(* Logix 5000 project; controller FV vendor 1 type 14 code 217 rev 31.11; software revision 31.00; part 2 of 63 *)

        [144]   // 0 0 0 min input
        [145]   // 0 0 0 max input
        [146]   // 0 0 0 min scaled
        [147]   // 0 0 0 max scale
        [148]   // 0 0 0 High Limit
        [149]   // 0 0 0 Low Limit
        [14]   // FV26/LTX01 FV26 level transmitter min input
        [151]   // 0 0 0 Flags
        [151].0   // 0 0 0 High
        [151].1   // 0 0 0 Low
        [151].15   // 0 0 0 Fault
        [152]   // 0 0 0 mA
        [153]   // 0 0 0 spare
        [154]   // 0 0 0 min input
        [155]   // 0 0 0 max input
        [156]   // 0 0 0 min scaled
        [157]   // 0 0 0 max scale
        [158]   // 0 0 0 High Limit
        [159]   // 0 0 0 Low Limit
        [15]   // FV26/LTX01 FV26 level transmitter max input
        [16]   // FV26/LTX01 FV26 level transmitter min scaled
        [17]   // FV26/LTX01 FV26 level transmitter max scale
        [18]   // FV26/LTX01 FV26 level transmitter High Limit
        [19]   // FV26/LTX01 FV26 level transmitter Low Limit
        [1]   // FV26/PTX01 FV26 top pressure Flags
        [1].0   // FV26/PTX01 FV26 top pressure High
        [1].1   // FV26/PTX01 FV26 top pressure Low
        [1].15   // FV26/PTX01 FV26 top pressure Fault
        [20]   // FV27/PTX01 FV27 top pressure transmitter
        [21]   // FV27/PTX01 FV27 top pressure Flags
        [21].0   // FV27/PTX01 FV27 top pressure High
        [21].1   // FV27/PTX01 FV27 top pressure Low
        [21].15   // FV27/PTX01 FV27 top pressure Fault
        [22]   // FV27/PTX01 FV27 top pressure mA
        [23]   // FV27/PTX01 FV27 top pressure spare
        [24]   // FV27/PTX01 FV27 top pressure min input
        [25]   // FV27/PTX01 FV27 top pressure max input
        [26]   // FV27/PTX01 FV27 top pressure min scaled
        [27]   // FV27/PTX01 FV27 top pressure max scale
        [28]   // FV27/PTX01 FV27 top pressure High Limit
        [29]   // FV27/PTX01 FV27 top pressure Low Limit
        [2]   // FV26/PTX01 FV26 top pressure mA
        [30]   // FV27/LTX01 FV27 level transmitter
        [31]   // FV27/LTX01 FV27 level transmitter Flags
        [31].0   // FV27/LTX01 FV27 level transmitter High
        [31].1   // FV27/LTX01 FV27 level transmitter Low
        [31].15   // FV27/LTX01 FV27 level transmitter Fault
        [32]   // FV27/LTX01 FV27 level transmitter mA
        [33]   // FV27/LTX01 FV27 level transmitter spare
        [34]   // FV27/LTX01 FV27 level transmitter min input
        [35]   // FV27/LTX01 FV27 level transmitter max input
        [36]   // FV27/LTX01 FV27 level transmitter min scaled
        [37]   // FV27/LTX01 FV27 level transmitter max scale
        [38]   // FV27/LTX01 FV27 level transmitter High Limit
        [39]   // FV27/LTX01 FV27 level transmitter Low Limit
        [3]   // FV26/PTX01 FV26 top pressure spare
        [40]   // FV28/PTX01 FV28 top pressure transmitter
        [41]   // FV28/PTX01 FV28 top pressure Flags
        [41].0   // FV28/PTX01 FV28 top pressure High
        [41].1   // FV28/PTX01 FV28 top pressure Low
        [41].15   // FV28/PTX01 FV28 top pressure Fault
        [42]   // FV28/PTX01 FV28 top pressure mA
        [43]   // FV28/PTX01 FV28 top pressure spare
        [44]   // FV28/PTX01 FV28 top pressure min input
        [45]   // FV28/PTX01 FV28 top pressure max input
        [46]   // FV28/PTX01 FV28 top pressure min scaled
        [47]   // FV28/PTX01 FV28 top pressure max scale
        [48]   // FV28/PTX01 FV28 top pressure High Limit
        [49]   // FV28/PTX01 FV28 top pressure Low Limit
        [4]   // FV26/PTX01 FV26 top pressure min input
        [50]   // FV28/LTX01 FV28 level transmitter
        [51]   // FV28/LTX01 FV28 level transmitter Flags
        [51].0   // FV28/LTX01 FV28 level transmitter High
        [51].1   // FV28/LTX01 FV28 level transmitter Low
        [51].15   // FV28/LTX01 FV28 level transmitter Fault
        [52]   // FV28/LTX01 FV28 level transmitter mA
        [53]   // FV28/LTX01 FV28 level transmitter spare
        [54]   // FV28/LTX01 FV28 level transmitter min input
        [55]   // FV28/LTX01 FV28 level transmitter max input
        [56]   // FV28/LTX01 FV28 level transmitter min scaled
        [57]   // FV28/LTX01 FV28 level transmitter max scale
        [58]   // FV28/LTX01 FV28 level transmitter High Limit
        [59]   // FV28/LTX01 FV28 level transmitter Low Limit
        [5]   // FV26/PTX01 FV26 top pressure max input
        [60]   // FV29/PTX01 FV29 top pressure transmitter
        [61]   // FV29/PTX01 FV29 top pressure Flags
        [61].0   // FV29/PTX01 FV29 top pressure High
        [61].1   // FV29/PTX01 FV29 top pressure Low
        [61].15   // FV29/PTX01 FV29 top pressure Fault
        [62]   // FV29/PTX01 FV29 top pressure mA
        [63]   // FV29/PTX01 FV29 top pressure spare
        [64]   // FV29/PTX01 FV29 top pressure min input
        [65]   // FV29/PTX01 FV29 top pressure max input
        [66]   // FV29/PTX01 FV29 top pressure min scaled
        [67]   // FV29/PTX01 FV29 top pressure max scale
        [68]   // FV29/PTX01 FV29 top pressure High Limit
        [69]   // FV29/PTX01 FV29 top pressure Low Limit
        [6]   // FV26/PTX01 FV26 top pressure min scaled
        [70]   // FV29/LTX01 FV29 level transmitter
        [71]   // FV29/LTX01 FV29 level transmitter Flags
        [71].0   // FV29/LTX01 FV29 level transmitter High
        [71].1   // FV29/LTX01 FV29 level transmitter Low
        [71].15   // FV29/LTX01 FV29 level transmitter Fault
        [72]   // FV29/LTX01 FV29 level transmitter mA
        [73]   // FV29/LTX01 FV29 level transmitter spare
        [74]   // FV29/LTX01 FV29 level transmitter min input
        [75]   // FV29/LTX01 FV29 level transmitter max input
        [76]   // FV29/LTX01 FV29 level transmitter min scaled
        [77]   // FV29/LTX01 FV29 level transmitter max scale
        [78]   // FV29/LTX01 FV29 level transmitter High Limit
        [79]   // FV29/LTX01 FV29 level transmitter Low Limit
        [7]   // FV26/PTX01 FV26 top pressure max scale
        [80]   // FV30/PTX01 FV30 top pressure transmitter
        [81]   // FV30/PTX01 FV30 top pressure Flags
        [81].0   // FV30/PTX01 FV30 top pressure High
        [81].1   // FV30/PTX01 FV30 top pressure Low
        [81].15   // FV30/PTX01 FV30 top pressure Fault
        [82]   // FV30/PTX01 FV30 top pressure mA
        [83]   // FV30/PTX01 FV30 top pressure spare
        [84]   // FV30/PTX01 FV30 top pressure min input
        [85]   // FV30/PTX01 FV30 top pressure max input
        [86]   // FV30/PTX01 FV30 top pressure min scaled
        [87]   // FV30/PTX01 FV30 top pressure max scale
        [88]   // FV30/PTX01 FV30 top pressure High Limit
        [89]   // FV30/PTX01 FV30 top pressure Low Limit
        [8]   // FV26/PTX01 FV26 top pressure High Limit
        [90]   // FV30/LTX01 FV30 level transmitter
        [91]   // FV30/LTX01 FV30 level transmitter Flags
        [91].0   // FV30/LTX01 FV30 level transmitter High
        [91].1   // FV30/LTX01 FV30 level transmitter Low
        [91].15   // FV30/LTX01 FV30 level transmitter Fault
        [92]   // FV30/LTX01 FV30 level transmitter mA
        [93]   // FV30/LTX01 FV30 level transmitter spare
        [94]   // FV30/LTX01 FV30 level transmitter min input
        [95]   // FV30/LTX01 FV30 level transmitter max input
        [96]   // FV30/LTX01 FV30 level transmitter min scaled
        [97]   // FV30/LTX01 FV30 level transmitter max scale
        [98]   // FV30/LTX01 FV30 level transmitter High Limit
        [99]   // FV30/LTX01 FV30 level transmitter Low Limit
        [9]   // FV26/PTX01 FV26 top pressure Low Limit
   FR_N201 : INT[265];   // Original N File From SLC, No Description Available
   FR_N207 : INT[265] := ([0] := 256, [1] := 1, [2] := 2, [3] := 3, [4] := 4, [5] := 5, [6] := 6, [7] := 7, [8] := 8, [9] := 9, [10] := 10, [11] := 11, [12] := 12, [13] := 13, [14] := 14, [15] := 15, [16] := 16, [17] := 17, [18] := 18, [19] := 19, [20] := 20, [21] := 21, [22] := 22, [23] := 23, [24] := 24, [25] := 25, [26] := 26, [27] := 27, [28] := 28, [29] := 29, [30] := 30, [31] := 31, [32] := 32, [33] := 33, [34] := 34, [35] := 35, [36] := 36, [37] := 37, [38] := 38, [39] := 39, [40] := 40, [41] := 41, [42] := 42, [43] := 43, [44] := 44, [45] := 45, [46] := 46, [47] := 47, [48] := 48, [49] := 49, [50] := 50, [51] := 51, [52] := 52, [53] := 53, [54] := 54, [55] := 55, [56] := 56, [57] := 57, [58] := 58, [59] := 59,
        [60] := 60, [61] := 61, [62] := 62, [63] := 63, [64] := 64, [65] := 65, [66] := 66, [67] := 67, [68] := 68, [69] := 69, [70] := 70, [71] := 71, [72] := 72, [73] := 73, [74] := 74, [75] := 75, [76] := 76, [77] := 77, [78] := 78, [79] := 79, [80] := 80, [81] := 81, [82] := 82, [83] := 83, [84] := 84, [85] := 85, [86] := 86, [87] := 87, [88] := 88, [89] := 89, [90] := 90, [91] := 91, [92] := 92, [93] := 93, [94] := 94, [95] := 95, [96] := 96, [97] := 97, [98] := 98, [99] := 99, [100] := 100, [101] := 101, [102] := 102, [103] := 103, [104] := 104, [105] := 105, [106] := 106, [107] := 107, [108] := 108, [109] := 109, [110] := 110, [111] := 111, [112] := 112, [113] := 113, [114] := 114, [115] := 115, [116] := 116, [117] := 117, [118] := 118, [119] := 119,
        [120] := 120, [121] := 121, [122] := 122, [123] := 123, [124] := 124, [125] := 125, [126] := 126, [127] := 127, [128] := 128, [129] := 129, [130] := 130, [131] := 131, [132] := 132, [133] := 133, [134] := 134, [135] := 135, [136] := 136, [137] := 137, [138] := 138, [139] := 139, [140] := 140, [141] := 141, [142] := 142, [143] := 143, [144] := 144, [145] := 145, [146] := 146, [147] := 147, [148] := 148, [149] := 149, [150] := 150, [151] := 151, [152] := 152, [153] := 153, [154] := 154, [155] := 155, [156] := 156, [157] := 157, [158] := 158, [159] := 159, [160] := 160, [161] := 161, [162] := 162, [163] := 163, [164] := 164, [165] := 165, [166] := 166, [167] := 167, [168] := 168, [169] := 169, [170] := 170, [171] := 171, [172] := 172, [173] := 173, [174] := 174, [175] := 175, [176] := 176, [177] := 177, [178] := 178, [179] := 179,
        [180] := 180, [181] := 181, [182] := 182, [183] := 183, [184] := 184, [185] := 185, [186] := 186, [187] := 187, [188] := 188, [189] := 189, [190] := 190, [191] := 191, [192] := 192, [193] := 193, [194] := 194, [195] := 195, [196] := 196, [197] := 197, [198] := 198, [199] := 199, [200] := 200, [201] := 201, [202] := 202, [203] := 203, [204] := 204, [205] := 205, [206] := 206, [207] := 207, [208] := 208, [209] := 209, [210] := 210, [211] := 211, [212] := 212, [213] := 213, [214] := 214, [215] := 215, [216] := 216, [217] := 217, [218] := 218, [219] := 219, [220] := 220, [221] := 221, [222] := 222, [223] := 223, [224] := 224, [225] := 225, [226] := 226, [227] := 227, [228] := 228, [229] := 229, [230] := 230, [231] := 231, [232] := 232, [233] := 233, [234] := 234, [235] := 235, [236] := 236, [237] := 237, [238] := 238, [239] := 239,
        [240] := 240, [241] := 241, [242] := 242, [243] := 243, [244] := 244, [245] := 245, [246] := 246, [247] := 247, [248] := 248, [249] := 249, [250] := 250, [251] := 251, [252] := 252, [253] := 253, [254] := 254, [255] := 255);   // Original N File From SLC, No Description Available
   FR_N21 : INT[265] := ([26] := 700, [27] := 700, [28] := 700, [29] := 700, [30] := 700, [31] := 700);   // CHASE_V FV Filling Beer Chas e Volumes
   FR_N210 : INT[265] := ([0] := 500, [1] := 12000, [2] := 18725, [5] := 1000, [6] := 4000, [7] := 20000, [8] := 6242, [9] := 31208, [11] := 12000, [12] := 18725, [15] := 1000, [16] := 4000, [17] := 20000, [18] := 6242, [19] := 31208, [20] := 500, [21] := 8800, [22] := 13732, [25] := 1000, [26] := 4000, [27] := 20000, [28] := 6242, [29] := 31208);   // ANALOG_OUT Analog Outputs
        [0]   // YM/P01 Yeast Main Pump 1 FV26-31 0.0-100.0%
        [10]   // YM/P02 Yeast Main Pump 2 FV1-17 0.0-100.0%
        [11]   // YM/P02 Yeast Main Pump 2 FV1-17 4.000-20.000mA
        [12]   // YM/P02 Yeast Main Pump 2 FV1-17 Output Card Scaling 6242-31209
        [1]   // YM/P01 Yeast Main Pump 1 FV26-31 4.000-20.000mA
        [20]   // YM/P03 Yeast Main Pump 3 FV18-25 0.0-100.0%
        [21]   // YM/P03 Yeast Main Pump 3 FV18-25 4.000-20.000mA
        [22]   // YM/P03 Yeast Main Pump 3 FV18-25 Output Card Scaling 6242-31210
        [2]   // YM/P01 Yeast Main Pump 1 FV26-31 Output Card Scaling 6242-31208
   FR_N220 : INT[265] := ([0] := 130, [1] := 110, [2] := -1, [3] := 5);   // CHECKLIST Checklist Loop Contr ollers
        [0]   // File containing Checklist
        [1]   // Pointer to item
        [2]   // Pointer to faulted item
        [3]   // Copy of Checkword Number
   FR_N225 : INT[265];   // Original N File From SLC, No Description Available
        [0].0   // Watchdog from GEA Tank Farm Both directions controlled by GEA
   FR_N226 : INT[265];   // Original N File From SLC, No Description Available
        [0].0   // Watchdog to GEA Tank Farm Both directions controlled by GEA
   FR_N245 : INT[265];   // CHECKWORD Checkword Loop Contr ol
        [0]   // Checkword Pointer
        [10].0   // Clear Manual, Reverse, Data & Fault Bits & Set Timer Presets to 30s
        [10].1   // Initialise Timers
        [11]   // Initialisation Pointer
        [12]   // Output OR Manual On
        [13].0   // Current item's output pointer OK
        [13].1   // Current item's energised input pointer OK
        [13].2   // Current item's deenergised input pointer OK
        [1]   // Current item's output pointer
        [21].1   // This Item is Reverse Acting i.e. Air to Close
        [21].2   // This Item is a Pump Energised bit is Run Feedback Deenergised bit is Tripped Signal
        [28]   // Number of items checked this scan
        [29]   // Number of items to check each scan
        [2]   // Current item's energised input pointer
        [3]   // Current item's deenergised input pointer
        [4]   // Current item's checkword
        [4].10   // Current item's checkword Energised Input
        [4].11   // Current item's checkword Deenergised Input
        [4].14   // Current Item Reverse Acting Flag
        [7]   // Current Item's Timer
        [9]   // Last Checkword Number
   FR_N252 : INT[265];   // OUTPUT_PTR Checkword Pointers t o output flags in B2 50
   FR_N253 : INT[265];   // EN_POINT Pointers to energise d input flags in B25 1
   FR_N254 : INT[265];   // DEN_POINT Pointers to deenergi sed input flags in B 251
   FR_N255 : INT[265] := ([0] := 2128, [1] := 2128, [2] := 2128, [3] := 2128, [4] := 2128, [5] := 2128, [6] := 2128, [7] := 10832, [8] := 1152, [9] := 2128, [10] := 2128, [11] := 2128, [12] := 2128, [13] := 1152, [14] := 2128, [15] := 2128, [16] := 2128, [17] := 2128, [18] := 2128, [19] := 2128, [20] := 2128, [21] := 2128, [22] := 2128, [23] := 2128, [24] := 2128, [25] := 1104, [26] := 2128, [27] := 1152, [28] := 2128, [29] := 2128, [30] := 2128, [31] := 2128, [32] := 1152, [33] := 2128, [34] := 2128, [35] := 2128, [36] := 2128, [37] := 2128, [38] := 2128, [39] := 2128, [40] := 1104, [41] := 2128, [42] := 2128, [43] := 2128, [44] := 1616, [45] := 2128, [46] := 2128, [47] := 2128, [48] := 2128, [49] := 2128, [50] := 2128, [51] := 2128, [52] := 2128, [53] := 2128, [54] := 2128, [55] := 2128, [56] := 2128, [57] := 2128, [58] := 2128, [59] := 2128,
        [60] := 2128, [61] := 2128, [62] := 2128, [63] := 2384, [64] := 1152, [65] := 2128, [66] := 2128, [67] := 2128, [68] := 2128, [69] := 1152, [70] := 2128, [71] := 2128, [72] := 2128, [73] := 2128, [74] := 2128, [75] := 2128, [76] := 2128, [77] := 1104, [78] := 2128, [79] := 2128, [84] := 2128, [85] := 2128, [86] := 2128, [87] := 2128, [88] := 2128, [89] := 2128, [90] := 2128, [91] := 1616, [92] := 1616, [93] := 2128, [94] := 2128, [95] := 2128, [96] := 2176, [97] := 2176, [98] := 2176, [99] := 2176, [100] := 2176, [101] := 2176);   // CHECKWORDS
        [0]   // FVS/P01 CIP return pump 0 Checkword CW0
        [0].13   // FVS/P01 CIP return pump 0 Inhibit Checking CW0
        [0].15   // FVS/P01 CIP return pump 0 Fault CW0
        [0].8   // FVS/P01 CIP return pump 0 Manual CW0
        [0].9   // FVS/P01 CIP return pump 0 Drive CW0
        [100].13   // FV30/AV08 FV30 Sprayball Inhibit Checking CW100
        [100].9   // FV30/AV08 FV30 Sprayball Drive CW100
        [101].13   // FV31/AV08 FV31 Sprayball Inhibit Checking CW101
        [101].9   // FV31/AV08 FV31 Sprayball Drive CW101
        [10]   // FV26/AV05 FV26 Green Beer 0 Checkword CW10
        [10].13   // FV26/AV05 FV26 Green Beer 0 Inhibit Checking CW10
        [10].15   // FV26/AV05 FV26 Green Beer 0 Fault CW10
        [10].8   // FV26/AV05 FV26 Green Beer 0 Manual CW10
        [10].9   // FV26/AV05 FV26 Green Beer 0 Drive CW10
        [11]   // FV26/AV06 FV26 Yeast Out 0 Checkword CW11
        [11].13   // FV26/AV06 FV26 Yeast Out 0 Inhibit Checking CW11
        [11].15   // FV26/AV06 FV26 Yeast Out 0 Fault CW11
        [11].8   // FV26/AV06 FV26 Yeast Out 0 Manual CW11
        [11].9   // FV26/AV06 FV26 Yeast Out 0 Drive CW11
        [12]   // FV26/AV07 FV26 CIP Return 0 Checkword CW12
        [12].13   // FV26/AV07 FV26 CIP Return 0 Inhibit Checking CW12
        [12].15   // FV26/AV07 FV26 CIP Return 0 Fault CW12
        [12].8   // FV26/AV07 FV26 CIP Return 0 Manual CW12
        [12].9   // FV26/AV07 FV26 CIP Return 0 Drive CW12
        [13]   // FV27/AV01 FV27 Filtrate Inlet 0 Checkword CW13
        [13].13   // FV27/AV01 FV27 Filtrate Inlet 0 Inhibit Checking CW13
        [13].14   // Reverse Acting
        [13].15   // FV27/AV01 FV27 Filtrate Inlet 0 Fault CW13
        [13].8   // FV27/AV01 FV27 Filtrate Inlet 0 Manual CW13
        [13].9   // FV27/AV01 FV27 Filtrate Inlet 0 Drive CW13
        [14]   // FV27/AV04 FV27 Filling 0 Checkword CW14
        [14].13   // FV27/AV04 FV27 Filling 0 Inhibit Checking CW14
        [14].15   // FV27/AV04 FV27 Filling 0 Fault CW14
        [14].8   // FV27/AV04 FV27 Filling 0 Manual CW14
        [14].9   // FV27/AV04 FV27 Filling 0 Drive CW14
        [15]   // FV27/AV05 FV27 Green Beer 0 Checkword CW15
        [15].13   // FV27/AV05 FV27 Green Beer 0 Inhibit Checking CW15
        [15].15   // FV27/AV05 FV27 Green Beer 0 Fault CW15
        [15].8   // FV27/AV05 FV27 Green Beer 0 Manual CW15
        [15].9   // FV27/AV05 FV27 Green Beer 0 Drive CW15
        [16]   // FV27/AV06 FV27 Yeast Out 0 Checkword CW16
        [16].13   // FV27/AV06 FV27 Yeast Out 0 Inhibit Checking CW16
        [16].15   // FV27/AV06 FV27 Yeast Out 0 Fault CW16
        [16].8   // FV27/AV06 FV27 Yeast Out 0 Manual CW16
        [16].9   // FV27/AV06 FV27 Yeast Out 0 Drive CW16
        [17]   // FV27/AV07 FV27 CIP Return 0 Checkword CW17
        [17].13   // FV27/AV07 FV27 CIP Return 0 Inhibit Checking CW17
        [17].15   // FV27/AV07 FV27 CIP Return 0 Fault CW17
        [17].8   // FV27/AV07 FV27 CIP Return 0 Manual CW17
        [17].9   // FV27/AV07 FV27 CIP Return 0 Drive CW17
        [18]   // VB1/AV01 VB1 Green Beer Main CIP Supply Checkword CW18
        [18].13   // VB1/AV01 VB1 Green Beer Main CIP Supply Inhibit Checking CW18
        [18].15   // VB1/AV01 VB1 Green Beer Main CIP Supply Fault CW18
        [18].8   // VB1/AV01 VB1 Green Beer Main CIP Supply Manual CW18
        [18].9   // VB1/AV01 VB1 Green Beer Main CIP Supply Drive CW18
        [19]   // VB1/AV02 VB1 Yeast Out Main CIP Supply Checkword CW19
        [19].13   // VB1/AV02 VB1 Yeast Out Main CIP Supply Inhibit Checking CW19
        [19].15   // VB1/AV02 VB1 Yeast Out Main CIP Supply Fault CW19
        [19].8   // VB1/AV02 VB1 Yeast Out Main CIP Supply Manual CW19
        [19].9   // VB1/AV02 VB1 Yeast Out Main CIP Supply Drive CW19
        [1]   // YM/P01 Yeast main (FV26-31) pump Checkword CW1
        [1].13   // YM/P01 Yeast main (FV26-31) pump Inhibit Checking CW1
        [1].15   // YM/P01 Yeast main (FV26-31) pump Fault CW1
        [1].8   // YM/P01 Yeast main (FV26-31) pump Manual CW1
        [1].9   // YM/P01 Yeast main (FV26-31) pump Drive CW1
        [20]   // VB1/AV03 VB1 Green Beer Main Water Chase Checkword CW20
        [20].13   // VB1/AV03 VB1 Green Beer Main Water Chase Inhibit Checking CW20
        [20].15   // VB1/AV03 VB1 Green Beer Main Water Chase Fault CW20
        [20].8   // VB1/AV03 VB1 Green Beer Main Water Chase Manual CW20
        [20].9   // VB1/AV03 VB1 Green Beer Main Water Chase Drive CW20
        [21]   // VB1/AV04 VB1 Yeast Out Main Water Chase Checkword CW21
        [21].13   // VB1/AV04 VB1 Yeast Out Main Water Chase Inhibit Checking CW21
        [21].15   // VB1/AV04 VB1 Yeast Out Main Water Chase Fault CW21
        [21].8   // VB1/AV04 VB1 Yeast Out Main Water Chase Manual CW21
        [21].9   // VB1/AV04 VB1 Yeast Out Main Water Chase Drive CW21
        [22]   // VB1/AV05 VB1 Filling Main Seat Clean Checkword CW22
        [22].13   // VB1/AV05 VB1 Filling Main Seat Clean Inhibit Checking CW22
        [22].15   // VB1/AV05 VB1 Filling Main Seat Clean Fault CW22
        [22].8   // VB1/AV05 VB1 Filling Main Seat Clean Manual CW22
        [22].9   // VB1/AV05 VB1 Filling Main Seat Clean Drive CW22
        [23]   // VB1/AV06 VB1 Green Beer Main Seat Clean Checkword CW23
        [23].13   // VB1/AV06 VB1 Green Beer Main Seat Clean Inhibit Checking CW23
        [23].15   // VB1/AV06 VB1 Green Beer Main Seat Clean Fault CW23
        [23].8   // VB1/AV06 VB1 Green Beer Main Seat Clean Manual CW23
        [23].9   // VB1/AV06 VB1 Green Beer Main Seat Clean Drive CW23
        [24]   // VB1/AV07 VB1 Yeast Out Main Seat Clean Checkword CW24
        [24].13   // VB1/AV07 VB1 Yeast Out Main Seat Clean Inhibit Checking CW24
        [24].15   // VB1/AV07 VB1 Yeast Out Main Seat Clean Fault CW24
        [24].8   // VB1/AV07 VB1 Yeast Out Main Seat Clean Manual CW24
        [24].9   // VB1/AV07 VB1 Yeast Out Main Seat Clean Drive CW24
        [25]   // VB1/AV08 VB1 Filling Main Block Checkword CW25
        [25].13   // VB1/AV08 VB1 Filling Main Block Inhibit Checking CW25
        [25].14   // Reverse Acting
        [25].15   // VB1/AV08 VB1 Filling Main Block Fault CW25
        [25].8   // VB1/AV08 VB1 Filling Main Block Manual CW25
        [25].9   // VB1/AV08 VB1 Filling Main Block Drive CW25
        [26]   // VB1/AV09 VB1 Filling Main Drain Checkword CW26
        [26].13   // VB1/AV09 VB1 Filling Main Drain Inhibit Checking CW26
        [26].15   // VB1/AV09 VB1 Filling Main Drain Fault CW26
        [26].8   // VB1/AV09 VB1 Filling Main Drain Manual CW26
        [26].9   // VB1/AV09 VB1 Filling Main Drain Drive CW26
        [27]   // FV28/AV01 FV28 Filtrate Inlet 0 Checkword CW27
        [27].13   // FV28/AV01 FV28 Filtrate Inlet 0 Inhibit Checking CW27
        [27].14   // Reverse Acting
        [27].15   // FV28/AV01 FV28 Filtrate Inlet 0 Fault CW27
        [27].8   // FV28/AV01 FV28 Filtrate Inlet 0 Manual CW27
        [27].9   // FV28/AV01 FV28 Filtrate Inlet 0 Drive CW27
        [28]   // FV28/AV04 FV28 Filling 0 Checkword CW28
        [28].13   // FV28/AV04 FV28 Filling 0 Inhibit Checking CW28
        [28].15   // FV28/AV04 FV28 Filling 0 Fault CW28
        [28].8   // FV28/AV04 FV28 Filling 0 Manual CW28
        [28].9   // FV28/AV04 FV28 Filling 0 Drive CW28
        [29]   // FV28/AV05 FV28 Green Beer 0 Checkword CW29
        [29].13   // FV28/AV05 FV28 Green Beer 0 Inhibit Checking CW29
        [29].15   // FV28/AV05 FV28 Green Beer 0 Fault CW29
        [29].8   // FV28/AV05 FV28 Green Beer 0 Manual CW29
        [29].9   // FV28/AV05 FV28 Green Beer 0 Drive CW29
        [2]   // GBM/P01 Green Beer main pump Checkword CW2
        [2].13   // GBM/P01 Green Beer main pump Inhibit Checking CW2
        [2].15   // GBM/P01 Green Beer main pump Fault CW2
        [2].8   // GBM/P01 Green Beer main pump Manual CW2
        [2].9   // GBM/P01 Green Beer main pump Drive CW2
        [30]   // FV28/AV06 FV28 Yeast Out 0 Checkword CW30
        [30].13   // FV28/AV06 FV28 Yeast Out 0 Inhibit Checking CW30
        [30].15   // FV28/AV06 FV28 Yeast Out 0 Fault CW30
        [30].8   // FV28/AV06 FV28 Yeast Out 0 Manual CW30
        [30].9   // FV28/AV06 FV28 Yeast Out 0 Drive CW30
        [31]   // FV28/AV07 FV28 CIP Return 0 Checkword CW31
        [31].13   // FV28/AV07 FV28 CIP Return 0 Inhibit Checking CW31
        [31].15   // FV28/AV07 FV28 CIP Return 0 Fault CW31
        [31].8   // FV28/AV07 FV28 CIP Return 0 Manual CW31
        [31].9   // FV28/AV07 FV28 CIP Return 0 Drive CW31
        [32]   // FV29/AV01 FV29 Filtrate Inlet 0 Checkword CW32
        [32].13   // FV29/AV01 FV29 Filtrate Inlet 0 Inhibit Checking CW32
        [32].14   // Reverse Acting
        [32].15   // FV29/AV01 FV29 Filtrate Inlet 0 Fault CW32
        [32].8   // FV29/AV01 FV29 Filtrate Inlet 0 Manual CW32
        [32].9   // FV29/AV01 FV29 Filtrate Inlet 0 Drive CW32
        [33]   // FV29/AV04 FV29 Filling 0 Checkword CW33
        [33].13   // FV29/AV04 FV29 Filling 0 Inhibit Checking CW33
        [33].15   // FV29/AV04 FV29 Filling 0 Fault CW33
        [33].8   // FV29/AV04 FV29 Filling 0 Manual CW33
        [33].9   // FV29/AV04 FV29 Filling 0 Drive CW33
        [34]   // FV29/AV05 FV29 Green Beer 0 Checkword CW34
        [34].13   // FV29/AV05 FV29 Green Beer 0 Inhibit Checking CW34
        [34].15   // FV29/AV05 FV29 Green Beer 0 Fault CW34
        [34].8   // FV29/AV05 FV29 Green Beer 0 Manual CW34
        [34].9   // FV29/AV05 FV29 Green Beer 0 Drive CW34
        [35]   // FV29/AV06 FV29 Yeast Out 0 Checkword CW35
        [35].13   // FV29/AV06 FV29 Yeast Out 0 Inhibit Checking CW35
        [35].15   // FV29/AV06 FV29 Yeast Out 0 Fault CW35
        [35].8   // FV29/AV06 FV29 Yeast Out 0 Manual CW35
        [35].9   // FV29/AV06 FV29 Yeast Out 0 Drive CW35
        [36]   // FV29/AV07 FV29 CIP Return 0 Checkword CW36
        [36].13   // FV29/AV07 FV29 CIP Return 0 Inhibit Checking CW36
        [36].15   // FV29/AV07 FV29 CIP Return 0 Fault CW36
        [36].8   // FV29/AV07 FV29 CIP Return 0 Manual CW36
        [36].9   // FV29/AV07 FV29 CIP Return 0 Drive CW36
        [37]   // VB2/AV01 VB2 Filling Main Seat Clean Checkword CW37
        [37].13   // VB2/AV01 VB2 Filling Main Seat Clean Inhibit Checking CW37
        [37].15   // VB2/AV01 VB2 Filling Main Seat Clean Fault CW37
        [37].8   // VB2/AV01 VB2 Filling Main Seat Clean Manual CW37
        [37].9   // VB2/AV01 VB2 Filling Main Seat Clean Drive CW37
        [38]   // VB2/AV02 VB2 Green Beer Main Seat Clean Checkword CW38
        [38].13   // VB2/AV02 VB2 Green Beer Main Seat Clean Inhibit Checking CW38
        [38].15   // VB2/AV02 VB2 Green Beer Main Seat Clean Fault CW38
        [38].8   // VB2/AV02 VB2 Green Beer Main Seat Clean Manual CW38
        [38].9   // VB2/AV02 VB2 Green Beer Main Seat Clean Drive CW38
        [39]   // VB2/AV03 VB2 Yeast Out Main Seat Clean Checkword CW39
        [39].13   // VB2/AV03 VB2 Yeast Out Main Seat Clean Inhibit Checking CW39
        [39].15   // VB2/AV03 VB2 Yeast Out Main Seat Clean Fault CW39
        [39].8   // VB2/AV03 VB2 Yeast Out Main Seat Clean Manual CW39
        [39].9   // VB2/AV03 VB2 Yeast Out Main Seat Clean Drive CW39
        [3]   // YM/P02 Yeast main (FV2) pump Checkword CW3
        [3].13   // YM/P02 Yeast main (FV2) pump Inhibit Checking CW3
        [3].15   // YM/P02 Yeast main (FV2) pump Fault CW3
        [3].8   // YM/P02 Yeast main (FV2) pump Manual CW3
        [3].9   // YM/P02 Yeast main (FV2) pump Drive CW3
        [40]   // VB2/AV04 VB2 Filling Main Block Checkword CW40
        [40].13   // VB2/AV04 VB2 Filling Main Block Inhibit Checking CW40
        [40].14   // Reverse Acting
        [40].15   // VB2/AV04 VB2 Filling Main Block Fault CW40
        [40].8   // VB2/AV04 VB2 Filling Main Block Manual CW40
        [40].9   // VB2/AV04 VB2 Filling Main Block Drive CW40
        [41]   // VB2/AV05 VB2 Filling Main Drain Checkword CW41
        [41].13   // VB2/AV05 VB2 Filling Main Drain Inhibit Checking CW41
        [41].15   // VB2/AV05 VB2 Filling Main Drain Fault CW41
        [41].8   // VB2/AV05 VB2 Filling Main Drain Manual CW41
        [41].9   // VB2/AV05 VB2 Filling Main Drain Drive CW41
        [42]   // VB4/AV01 VB4 FV26 Vent Checkword CW42
        [42].13   // VB4/AV01 VB4 FV26 Vent Inhibit Checking CW42
        [42].15   // VB4/AV01 VB4 FV26 Vent Fault CW42
        [42].8   // VB4/AV01 VB4 FV26 Vent Manual CW42
        [42].9   // VB4/AV01 VB4 FV26 Vent Drive CW42
        [43]   // VB4/AV02 VB4 FV27 Vent Checkword CW43
        [43].13   // VB4/AV02 VB4 FV27 Vent Inhibit Checking CW43
        [43].15   // VB4/AV02 VB4 FV27 Vent Fault CW43
        [43].8   // VB4/AV02 VB4 FV27 Vent Manual CW43
        [43].9   // VB4/AV02 VB4 FV27 Vent Drive CW43
        [44]   // VB4/AV03 VB4 FV31 Vent Checkword CW44
        [44].13   // VB4/AV03 VB4 FV31 Vent Inhibit Checking CW44
        [44].15   // VB4/AV03 VB4 FV31 Vent Fault CW44
        [44].8   // VB4/AV03 VB4 FV31 Vent Manual CW44
        [44].9   // VB4/AV03 VB4 FV31 Vent Drive CW44
        [45]   // VB4/AV04 VB4 FV30 Vent Checkword CW45
        [45].13   // VB4/AV04 VB4 FV30 Vent Inhibit Checking CW45
        [45].15   // VB4/AV04 VB4 FV30 Vent Fault CW45
        [45].8   // VB4/AV04 VB4 FV30 Vent Manual CW45
        [45].9   // VB4/AV04 VB4 FV30 Vent Drive CW45
        [46]   // VB4/AV05 VB4 FV29 Vent Checkword CW46
        [46].13   // VB4/AV05 VB4 FV29 Vent Inhibit Checking CW46
        [46].15   // VB4/AV05 VB4 FV29 Vent Fault CW46
        [46].8   // VB4/AV05 VB4 FV29 Vent Manual CW46
        [46].9   // VB4/AV05 VB4 FV29 Vent Drive CW46
        [47]   // VB4/AV06 VB4 FV28 Vent Checkword CW47
        [47].13   // VB4/AV06 VB4 FV28 Vent Inhibit Checking CW47
        [47].15   // VB4/AV06 VB4 FV28 Vent Fault CW47
        [47].8   // VB4/AV06 VB4 FV28 Vent Manual CW47
        [47].9   // VB4/AV06 VB4 FV28 Vent Drive CW47
        [48]   // VB4/AV07 VB4 FV26 CIP Supply Checkword CW48
        [48].13   // VB4/AV07 VB4 FV26 CIP Supply Inhibit Checking CW48
        [48].15   // VB4/AV07 VB4 FV26 CIP Supply Fault CW48
        [48].8   // VB4/AV07 VB4 FV26 CIP Supply Manual CW48
        [48].9   // VB4/AV07 VB4 FV26 CIP Supply Drive CW48
        [49]   // VB4/AV08 VB4 FV27 CIP Supply Checkword CW49
        [49].13   // VB4/AV08 VB4 FV27 CIP Supply Inhibit Checking CW49
        [49].15   // VB4/AV08 VB4 FV27 CIP Supply Fault CW49
        [49].8   // VB4/AV08 VB4 FV27 CIP Supply Manual CW49
        [49].9   // VB4/AV08 VB4 FV27 CIP Supply Drive CW49
        [4]   // YM/P03 Yeast main (FV18-25) pump Checkword CW4
        [4].13   // YM/P03 Yeast main (FV18-25) pump Inhibit Checking CW4
        [4].15   // YM/P03 Yeast main (FV18-25) pump Fault CW4
        [4].8   // YM/P03 Yeast main (FV18-25) pump Manual CW4
        [4].9   // YM/P03 Yeast main (FV18-25) pump Drive CW4
        [50]   // VB4/AV09 VB4 FV31 CIP Supply Checkword CW50
        [50].13   // VB4/AV09 VB4 FV31 CIP Supply Inhibit Checking CW50
        [50].15   // VB4/AV09 VB4 FV31 CIP Supply Fault CW50
        [50].8   // VB4/AV09 VB4 FV31 CIP Supply Manual CW50
        [50].9   // VB4/AV09 VB4 FV31 CIP Supply Drive CW50
        [51]   // VB4/AV10 VB4 FV30 CIP Supply Checkword CW51
        [51].13   // VB4/AV10 VB4 FV30 CIP Supply Inhibit Checking CW51
        [51].15   // VB4/AV10 VB4 FV30 CIP Supply Fault CW51
        [51].8   // VB4/AV10 VB4 FV30 CIP Supply Manual CW51
        [51].9   // VB4/AV10 VB4 FV30 CIP Supply Drive CW51
        [52]   // VB4/AV11 VB4 FV29 CIP Supply Checkword CW52
        [52].13   // VB4/AV11 VB4 FV29 CIP Supply Inhibit Checking CW52
        [52].15   // VB4/AV11 VB4 FV29 CIP Supply Fault CW52
        [52].8   // VB4/AV11 VB4 FV29 CIP Supply Manual CW52
        [52].9   // VB4/AV11 VB4 FV29 CIP Supply Drive CW52
        [53]   // VB4/AV12 VB4 FV28 CIP Supply Checkword CW53
        [53].13   // VB4/AV12 VB4 FV28 CIP Supply Inhibit Checking CW53
        [53].15   // VB4/AV12 VB4 FV28 CIP Supply Fault CW53
        [53].8   // VB4/AV12 VB4 FV28 CIP Supply Manual CW53
        [53].9   // VB4/AV12 VB4 FV28 CIP Supply Drive CW53
        [54]   // VB4/AV13 VB4 FV26 Filtrate Supply Checkword CW54
        [54].13   // VB4/AV13 VB4 FV26 Filtrate Supply Inhibit Checking CW54
        [54].15   // VB4/AV13 VB4 FV26 Filtrate Supply Fault CW54
        [54].8   // VB4/AV13 VB4 FV26 Filtrate Supply Manual CW54
        [54].9   // VB4/AV13 VB4 FV26 Filtrate Supply Drive CW54
        [55]   // VB4/AV14 VB4 FV27 Filtrate Supply Checkword CW55
        [55].13   // VB4/AV14 VB4 FV27 Filtrate Supply Inhibit Checking CW55
        [55].15   // VB4/AV14 VB4 FV27 Filtrate Supply Fault CW55
        [55].8   // VB4/AV14 VB4 FV27 Filtrate Supply Manual CW55
        [55].9   // VB4/AV14 VB4 FV27 Filtrate Supply Drive CW55
        [56]   // VB4/AV15 VB4 FV31 Filtrate Supply Checkword CW56
        [56].13   // VB4/AV15 VB4 FV31 Filtrate Supply Inhibit Checking CW56
        [56].15   // VB4/AV15 VB4 FV31 Filtrate Supply Fault CW56
        [56].8   // VB4/AV15 VB4 FV31 Filtrate Supply Manual CW56
        [56].9   // VB4/AV15 VB4 FV31 Filtrate Supply Drive CW56
        [57]   // VB4/AV23 VB4 Filtrate Drain 0 Checkword CW57
        [57].13   // VB4/AV23 VB4 Filtrate Drain 0 Inhibit Checking CW57
        [57].15   // VB4/AV23 VB4 Filtrate Drain 0 Fault CW57
        [57].8   // VB4/AV23 VB4 Filtrate Drain 0 Manual CW57
        [57].9   // VB4/AV23 VB4 Filtrate Drain 0 Drive CW57
        [58]   // VB4/AV17 VB4 FV29 Filtrate Supply Checkword CW58
        [58].13   // VB4/AV17 VB4 FV29 Filtrate Supply Inhibit Checking CW58
        [58].15   // VB4/AV17 VB4 FV29 Filtrate Supply Fault CW58
        [58].8   // VB4/AV17 VB4 FV29 Filtrate Supply Manual CW58
        [58].9   // VB4/AV17 VB4 FV29 Filtrate Supply Drive CW58
        [59]   // VB4/AV18 VB4 FV28 Filtrate Supply Checkword CW59
        [59].13   // VB4/AV18 VB4 FV28 Filtrate Supply Inhibit Checking CW59
        [59].15   // VB4/AV18 VB4 FV28 Filtrate Supply Fault CW59
        [59].8   // VB4/AV18 VB4 FV28 Filtrate Supply Manual CW59
        [59].9   // VB4/AV18 VB4 FV28 Filtrate Supply Drive CW59
        [5]   // FVR1/P01 Filtrate return pump Checkword CW5
        [5].13   // FVR1/P01 Filtrate return pump Inhibit Checking CW5
        [5].15   // FVR1/P01 Filtrate return pump Fault CW5
        [5].8   // FVR1/P01 Filtrate return pump Manual CW5
        [5].9   // FVR1/P01 Filtrate return pump Drive CW5
        [60]   // VB4/AV19 VB4 Filtrate Supply CIP Return Checkword CW60
        [60].13   // VB4/AV19 VB4 Filtrate Supply CIP Return Inhibit Checking CW60
        [60].15   // VB4/AV19 VB4 Filtrate Supply CIP Return Fault CW60
        [60].8   // VB4/AV19 VB4 Filtrate Supply CIP Return Manual CW60
        [60].9   // VB4/AV19 VB4 Filtrate Supply CIP Return Drive CW60
        [61]   // VB4/AV20 VB4 CIP Supply Seat Clean Checkword CW61
        [61].13   // VB4/AV20 VB4 CIP Supply Seat Clean Inhibit Checking CW61
        [61].15   // VB4/AV20 VB4 CIP Supply Seat Clean Fault CW61
        [61].8   // VB4/AV20 VB4 CIP Supply Seat Clean Manual CW61
        [61].9   // VB4/AV20 VB4 CIP Supply Seat Clean Drive CW61
        [62]   // VB4/AV21 VB4 Filtrate Supply Seat Clean Checkword CW62
        [62].13   // VB4/AV21 VB4 Filtrate Supply Seat Clean Inhibit Checking CW62
        [62].15   // VB4/AV21 VB4 Filtrate Supply Seat Clean Fault CW62
        [62].8   // VB4/AV21 VB4 Filtrate Supply Seat Clean Manual CW62
        [62].9   // VB4/AV21 VB4 Filtrate Supply Seat Clean Drive CW62
        [63]   // VB4/AV22 VB4 Vent Drain 0 Checkword CW63
        [63].13   // VB4/AV22 VB4 Vent Drain 0 Inhibit Checking CW63
        [63].15   // VB4/AV22 VB4 Vent Drain 0 Fault CW63
        [63].8   // VB4/AV22 VB4 Vent Drain 0 Manual CW63
        [63].9   // VB4/AV22 VB4 Vent Drain 0 Drive CW63
        [64]   // FV30/AV01 FV30 Filtrate Inlet 0 Checkword CW64
        [64].13   // FV30/AV01 FV30 Filtrate Inlet 0 Inhibit Checking CW64
        [64].14   // FV30/AV01 FV30 Filtrate Inlet 0 Reverse Acting CW64
        [64].15   // FV30/AV01 FV30 Filtrate Inlet 0 Fault CW64
        [64].8   // FV30/AV01 FV30 Filtrate Inlet 0 Manual CW64
        [64].9   // FV30/AV01 FV30 Filtrate Inlet 0 Drive CW64
        [65]   // FV30/AV04 FV30 Filling 0 Checkword CW65
        [65].13   // FV30/AV04 FV30 Filling 0 Inhibit Checking CW65
        [65].15   // FV30/AV04 FV30 Filling 0 Fault CW65
        [65].8   // FV30/AV04 FV30 Filling 0 Manual CW65
        [65].9   // FV30/AV04 FV30 Filling 0 Drive CW65
        [66]   // FV30/AV05 FV30 Green Beer 0 Checkword CW66
        [66].13   // FV30/AV05 FV30 Green Beer 0 Inhibit Checking CW66
        [66].15   // FV30/AV05 FV30 Green Beer 0 Fault CW66
        [66].8   // FV30/AV05 FV30 Green Beer 0 Manual CW66
        [66].9   // FV30/AV05 FV30 Green Beer 0 Drive CW66
        [67]   // FV30/AV06 FV30 Yeast Out 0 Checkword CW67
        [67].13   // FV30/AV06 FV30 Yeast Out 0 Inhibit Checking CW67
        [67].15   // FV30/AV06 FV30 Yeast Out 0 Fault CW67
        [67].8   // FV30/AV06 FV30 Yeast Out 0 Manual CW67
        [67].9   // FV30/AV06 FV30 Yeast Out 0 Drive CW67
        [68]   // FV30/AV07 FV30 CIP Return 0 Checkword CW68
        [68].13   // FV30/AV07 FV30 CIP Return 0 Inhibit Checking CW68
        [68].15   // FV30/AV07 FV30 CIP Return 0 Fault CW68
        [68].8   // FV30/AV07 FV30 CIP Return 0 Manual CW68
        [68].9   // FV30/AV07 FV30 CIP Return 0 Drive CW68
        [69]   // FV31/AV01 FV31 Filtrate Inlet 0 Checkword CW69
        [69].13   // FV31/AV01 FV31 Filtrate Inlet 0 Inhibit Checking CW69
        [69].14   // FV31/AV01 FV31 Filtrate Inlet 0 Reverse ACting CW69
        [69].15   // FV31/AV01 FV31 Filtrate Inlet 0 Fault CW69
        [69].8   // FV31/AV01 FV31 Filtrate Inlet 0 Manual CW69
        [69].9   // FV31/AV01 FV31 Filtrate Inlet 0 Drive CW69
        [6]   // 0 0 0 Checkword CW6
        [6].13   // 0 0 0 Inhibit Checking CW6
        [6].15   // 0 0 0 Fault CW6
        [6].8   // 0 0 0 Manual CW6
        [6].9   // 0 0 0 Drive CW6
        [70]   // FV31/AV04 FV31 Filling 0 Checkword CW70
        [70].13   // FV31/AV04 FV31 Filling 0 Inhibit Checking CW70
        [70].15   // FV31/AV04 FV31 Filling 0 Fault CW70
        [70].8   // FV31/AV04 FV31 Filling 0 Manual CW70
        [70].9   // FV31/AV04 FV31 Filling 0 Drive CW70
        [71]   // FV31/AV05 FV31 Green Beer 0 Checkword CW71
        [71].13   // FV31/AV05 FV31 Green Beer 0 Inhibit Checking CW71
        [71].15   // FV31/AV05 FV31 Green Beer 0 Fault CW71
        [71].8   // FV31/AV05 FV31 Green Beer 0 Manual CW71
        [71].9   // FV31/AV05 FV31 Green Beer 0 Drive CW71
        [72]   // FV31/AV06 FV31 Yeast Out 0 Checkword CW72
        [72].13   // FV31/AV06 FV31 Yeast Out 0 Inhibit Checking CW72
        [72].15   // FV31/AV06 FV31 Yeast Out 0 Fault CW72
        [72].8   // FV31/AV06 FV31 Yeast Out 0 Manual CW72
        [72].9   // FV31/AV06 FV31 Yeast Out 0 Drive CW72
        [73]   // FV31/AV07 FV31 CIP Return 0 Checkword CW73
        [73].13   // FV31/AV07 FV31 CIP Return 0 Inhibit Checking CW73
        [73].15   // FV31/AV07 FV31 CIP Return 0 Fault CW73
        [73].8   // FV31/AV07 FV31 CIP Return 0 Manual CW73
        [73].9   // FV31/AV07 FV31 CIP Return 0 Drive CW73
        [74]   // VB3/AV01 VB3 Filling Main Seat Clean Checkword CW74
        [74].13   // VB3/AV01 VB3 Filling Main Seat Clean Inhibit Checking CW74
        [74].15   // VB3/AV01 VB3 Filling Main Seat Clean Fault CW74
        [74].8   // VB3/AV01 VB3 Filling Main Seat Clean Manual CW74
        [74].9   // VB3/AV01 VB3 Filling Main Seat Clean Drive CW74
        [75]   // VB3/AV02 VB3 Green Beer Main Seat Clean Checkword CW75
        [75].13   // VB3/AV02 VB3 Green Beer Main Seat Clean Inhibit Checking CW75
        [75].15   // VB3/AV02 VB3 Green Beer Main Seat Clean Fault CW75
        [75].8   // VB3/AV02 VB3 Green Beer Main Seat Clean Manual CW75
        [75].9   // VB3/AV02 VB3 Green Beer Main Seat Clean Drive CW75
        [76]   // VB3/AV03 VB3 Yeast Out Main Seat Clean Checkword CW76
        [76].13   // VB3/AV03 VB3 Yeast Out Main Seat Clean Inhibit Checking CW76
        [76].15   // VB3/AV03 VB3 Yeast Out Main Seat Clean Fault CW76
        [76].8   // VB3/AV03 VB3 Yeast Out Main Seat Clean Manual CW76
        [76].9   // VB3/AV03 VB3 Yeast Out Main Seat Clean Drive CW76
        [77]   // VB3/AV04 VB3 Filling Main Block Checkword CW77
        [77].13   // VB3/AV04 VB3 Filling Main Block Inhibit Checking CW77
        [77].15   // VB3/AV04 VB3 Filling Main Block Fault CW77
        [77].8   // VB3/AV04 VB3 Filling Main Block Manual CW77
        [77].9   // VB3/AV04 VB3 Filling Main Block Drive CW77
        [78]   // VB3/AV05 VB3 Filling Main Drain Checkword CW78
        [78].13   // VB3/AV05 VB3 Filling Main Drain Inhibit Checking CW78
        [78].15   // VB3/AV05 VB3 Filling Main Drain Fault CW78
        [78].8   // VB3/AV05 VB3 Filling Main Drain Manual CW78
        [78].9   // VB3/AV05 VB3 Filling Main Drain Drive CW78
        [79]   // VB4/AV16 VB4 FV30 Filtrate Supply Checkword CW79
        [79].13   // VB4/AV16 VB4 FV30 Filtrate Supply Inhibit Checking CW79
        [79].15   // VB4/AV16 VB4 FV30 Filtrate Supply Fault CW79
        [79].8   // VB4/AV16 VB4 FV30 Filtrate Supply Manual CW79
        [79].9   // VB4/AV16 VB4 FV30 Filtrate Supply Drive CW79
        [7]   // FRV/AV01 Filtrate return Valve Checkword CW7
        [7].13   // FRV/AV01 Filtrate return Valve Inhibit Checking CW7
        [7].15   // FRV/AV01 Filtrate return Valve Fault CW7
        [7].8   // FRV/AV01 Filtrate return Valve Manual CW7
        [7].9   // FRV/AV01 Filtrate return Valve Drive CW7
        [80]   // 0 0 0 Checkword CW80
        [80].13   // 0 0 0 Inhibit Checking CW80
        [80].15   // 0 0 0 Fault CW80
        [80].8   // 0 0 0 Manual CW80
        [80].9   // 0 0 0 Drive CW80
        [81]   // 0 0 0 Checkword CW81
        [81].13   // 0 0 0 Inhibit Checking CW81
        [81].15   // 0 0 0 Fault CW81
        [81].8   // 0 0 0 Manual CW81
        [81].9   // 0 0 0 Drive CW81
        [82]   // 0 0 0 Checkword CW82
        [82].13   // 0 0 0 Inhibit Checking CW82
        [82].15   // 0 0 0 Fault CW82
        [82].8   // 0 0 0 Manual CW82
        [82].9   // 0 0 0 Drive CW82
        [83]   // 0 0 0 Checkword CW83
        [83].13   // 0 0 0 Inhibit Checking CW83
        [83].15   // 0 0 0 Fault CW83
        [83].8   // 0 0 0 Manual CW83
        [83].9   // 0 0 0 Drive CW83
        [84]   // 0 0 0 Checkword CW84
        [84].13   // 0 0 0 Inhibit Checking CW84
        [84].15   // 0 0 0 Fault CW84
        [84].8   // 0 0 0 Manual CW84
        [84].9   // 0 0 0 Drive CW84
        [85]   // 0 0 0 Checkword CW85
        [85].13   // 0 0 0 Inhibit Checking CW85
        [85].15   // 0 0 0 Fault CW85
        [85].8   // 0 0 0 Manual CW85
        [85].9   // 0 0 0 Drive CW85
        [86]   // 0 0 0 Checkword CW86
        [86].13   // 0 0 0 Inhibit Checking CW86
        [86].15   // 0 0 0 Fault CW86
        [86].8   // 0 0 0 Manual CW86
        [86].9   // 0 0 0 Drive CW86
        [87]   // 0 0 0 Checkword CW87
        [87].13   // 0 0 0 Inhibit Checking CW87
        [87].15   // 0 0 0 Fault CW87
        [87].8   // 0 0 0 Manual CW87
        [87].9   // 0 0 0 Drive CW87
        [88]   // FV26/VA01 FV26 vent actuator 0 Checkword CW88
        [88].13   // FV26/VA01 FV26 vent actuator 0 Inhibit Checking CW88
        [88].15   // FV26/VA01 FV26 vent actuator 0 Fault CW88
        [88].8   // FV26/VA01 FV26 vent actuator 0 Manual CW88
        [88].9   // FV26/VA01 FV26 vent actuator 0 Drive CW88
        [89]   // FV27/VA01 FV27 vent actuator 0 Checkword CW89
        [89].13   // FV27/VA01 FV27 vent actuator 0 Inhibit Checking CW89
        [89].15   // FV27/VA01 FV27 vent actuator 0 Fault CW89
        [89].8   // FV27/VA01 FV27 vent actuator 0 Manual CW89
        [89].9   // FV27/VA01 FV27 vent actuator 0 Drive CW89
        [8]   // FV26/AV01 FV26 Filtrate Inlet 0 Checkword CW8
        [8].13   // FV26/AV01 FV26 Filtrate Inlet 0 Inhibit Checking CW8
        [8].14   // Reverse Acting
        [8].15   // FV26/AV01 FV26 Filtrate Inlet 0 Fault CW8
        [8].8   // FV26/AV01 FV26 Filtrate Inlet 0 Manual CW8
        [8].9   // FV26/AV01 FV26 Filtrate Inlet 0 Drive CW8
        [90]   // FV28/VA01 FV28 vent actuator 0 Checkword CW90
        [90].13   // FV28/VA01 FV28 vent actuator 0 Inhibit Checking CW90
        [90].15   // FV28/VA01 FV28 vent actuator 0 Fault CW90
        [90].8   // FV28/VA01 FV28 vent actuator 0 Manual CW90
        [90].9   // FV28/VA01 FV28 vent actuator 0 Drive CW90
        [91]   // FV29/VA01 FV29 vent actuator 0 Checkword CW91
        [91].13   // FV29/VA01 FV29 vent actuator 0 Inhibit Checking CW91
        [91].15   // FV29/VA01 FV29 vent actuator 0 Fault CW91
        [91].8   // FV29/VA01 FV29 vent actuator 0 Manual CW91
        [91].9   // FV29/VA01 FV29 vent actuator 0 Drive CW91
        [92]   // FV30/VA01 FV30 vent actuator 0 Checkword CW92
        [92].13   // FV30/VA01 FV30 vent actuator 0 Inhibit Checking CW92
        [92].15   // FV30/VA01 FV30 vent actuator 0 Fault CW92
        [92].8   // FV30/VA01 FV30 vent actuator 0 Manual CW92
        [92].9   // FV30/VA01 FV30 vent actuator 0 Drive CW92
        [93]   // FV31/VA01 FV31 vent actuator 0 Checkword CW93
        [93].13   // FV31/VA01 FV31 vent actuator 0 Inhibit Checking CW93
        [93].15   // FV31/VA01 FV31 vent actuator 0 Fault CW93
        [93].8   // FV31/VA01 FV31 vent actuator 0 Manual CW93
        [93].9   // FV31/VA01 FV31 vent actuator 0 Drive CW93
        [94]   // AUDI1 CIP circulating audible alarm Checkword CW94
        [94].13   // AUDI1 CIP circulating audible alarm Inhibit Checking CW94
        [94].15   // AUDI1 CIP circulating audible alarm Fault CW94
        [94].8   // AUDI1 CIP circulating audible alarm Manual CW94
        [94].9   // AUDI1 CIP circulating audible alarm Drive CW94
        [95]   // BEACON1 CIP circulating flashing alarm Checkword CW95
        [95].13   // BEACON1 CIP circulating flashing alarm Inhibit Checking CW95
        [95].15   // BEACON1 CIP circulating flashing alarm Fault CW95
        [95].8   // BEACON1 CIP circulating flashing alarm Manual CW95
        [95].9   // BEACON1 CIP circulating flashing alarm Drive CW95
        [96].13   // FV26/AV08 FV26 Sprayball Inhibit Checking CW96
        [96].9   // FV26/AV08 FV26 Sprayball Drive CW96
        [97].13   // FV27/AV08 FV27 Sprayball Inhibit Checking CW97
        [97].9   // FV27/AV08 FV27 Sprayball Drive CW97
        [98].13   // FV28/AV08 FV28 Sprayball Inhibit Checking CW98
        [98].9   // FV28/AV08 FV28 Sprayball Drive CW98
        [99].13   // FV29/AV08 FV29 Sprayball Inhibit Checking CW99
        [99].9   // FV29/AV08 FV29 Sprayball Drive CW99
        [9]   // FV26/AV04 FV26 Filling 0 Checkword CW9
        [9].13   // FV26/AV04 FV26 Filling 0 Inhibit Checking CW9
        [9].15   // FV26/AV04 FV26 Filling 0 Fault CW9
        [9].8   // FV26/AV04 FV26 Filling 0 Manual CW9
        [9].9   // FV26/AV04 FV26 Filling 0 Drive CW9
   FR_N26 : INT[265] := ([0] := 226, [1] := 2, [3] := 1, [4] := 20, [5] := 1, [6] := 8, [7] := 1, [8] := 13226, [9] := -1, [10] := 669, [11] := 5336, [12] := 1575, [13] := 2902, [14] := 265, [15] := 667, [16] := 460, [17] := 4689, [18] := 12, [19] := 4633, [20] := 1, [21] := 21, [22] := -125, [23] := 50, [24] := -75, [25] := -175, [26] := 1000, [27] := 8, [30] := 20, [33] := 1, [37] := 702, [38] := 667, [52] := 1, [60] := 2, [68] := 2487, [69] := 2487, [100] := 42, [101] := 48, [102] := 54, [103] := 8, [104] := 9, [105] := 10, [106] := 11, [107] := 12, [108] := 96, [109] := -1, [110] := -1, [111] := -1, [112] := -1, [113] := -1, [114] := -1, [115] := -1, [116] := -1, [117] := -1, [118] := -1, [119] := -1, [120] := -1, [121] := -1, [122] := -1, [123] := -1, [124] := -1,
        [125] := -1, [126] := -1, [127] := -1, [128] := -1, [129] := -1, [130] := -1, [131] := -1, [132] := -1, [133] := -1, [134] := -1, [135] := -1, [136] := -1, [137] := -1, [138] := -1, [139] := -1, [140] := -1, [141] := -1, [142] := -1, [143] := -1, [144] := -1, [145] := -1, [146] := -1, [147] := -1, [148] := -1, [149] := -1);   // FV26
        [0]   // FV26
        [100]   // FV26 Checklist Data
        [10]   // FV26 Bottom Pressure
        [11]   // FV26 Damped Level
        [12]   // FV26 Cone Radius
        [13]   // FV26 Cone Height Estimate _ Probe not at bottom of vessel
        [14]   // FV26 Volume (HL)
        [19]   // FV26 Height above LTX
        [1]   // FV26 Status 0=Clean,1=Fill,2=Par t,3=Ferment,4=?,5=?, 6=?,7=?,8=Emptying,9 =Dirty,10-13=CIP
        [20]   // FV26 Top Pressure Bits
        [20].2   // FV26 Top Pressure Chill Down
        [20].5   // FV26 Top Pressure Step Channel 1 CIP
        [20].6   // FV26 Top Pressure Bits Ch1 CIP Complete
        [20].7   // FV26 Top Pressure Step Channel 2 CIP
        [20].8   // FV26 Top Pressure Bits Ch2 CIP Complete
        [21]   // FV26 Top Pressure Step Flags
        [21].0   // FV26 Top Pressure Control Over Pressure
        [21].12   // FV26 CIP Drain Down
        [21].4   // FV26 Top Pressure Open Vent
        [21].5   // FV26 Top Pressure Control Open Vent Actuator
        [21].6   // FV26 Over Top Pressure Limit
        [21].8   // FV26 Top Pressure Control Over Pressure Alarm
        [22]   // FV26 Top Pressure Setpoint
        [23]   // FV26 Top Pressure Deadband
        [24]   // FV26 Top Pressure Upper Limit
        [25]   // FV26 Top Pressure Lower Limit
        [26]   // FV26 Fermenting Pressure
        [27]   // FV26 Chill Down Time